DATA_BLOCK "DB_M256M_Scada"   // DB2011
{ S7_Optimized_Access := 'FALSE' }
VERSION : 0.1
   VAR
      tAlm : Struct   // HMI Alarms
         tE : Struct
            x0 : Bool;   // KE.Main emergency on
            x1 : Bool;   // KE1.Local emergency on
            x2 : Bool;   // Cabinet.Emergency localization
            x3 : Bool;   // SB1.Emergency localization
            x4 : Bool;   // SB2.Emergency localization
            x5 : Bool;
            x6 : Bool;
            x7 : Bool;
            x8 : Bool;
            x9 : Bool;
            x10 : Bool;
            x11 : Bool;
            x12 : Bool;
            x13 : Bool;
            x14 : Bool;
            x15 : Bool;
            x16 : Bool;
            x17 : Bool;
            x18 : Bool;
            x19 : Bool;
            x20 : Bool;
            x21 : Bool;
            x22 : Bool;
            x23 : Bool;
            x24 : Bool;
            x25 : Bool;
            x26 : Bool;
            x27 : Bool;
            x28 : Bool;
            x29 : Bool;
            x30 : Bool;
            x31 : Bool;
         END_STRUCT;
         tS : Struct
            tS0 : Struct
               x0 : Bool;   // xB18-3L+.PowerSupplyInputControlCabinetON / Head#1.Initialization timeout
               x1 : Bool;   // xB140QF2.ProtectionPowerSupplyMotorsYcut" / Head#1.homing timeout
               x2 : Bool;   // PLCA.Timeout receiving consumed message / Head#1.positioning timeout
               x3 : Bool;   // Syncro.Timeout receiving meter signal from main line / Head#1.carriage overload
               x4 : Bool;   // Head#1.drive error
               x5 : Bool;   // Head#1.missing ethernet IP connection
               x6 : Bool;   // Head#1.op.side overstroke
               x7 : Bool;   // Head#1.oppo.op.side overstroke
               x8 : Bool;   // Head#1.overstroke
               x9 : Bool;   // xB18-7L+.InputInstallationPowerSupplyON" / Head#2.Initialization timeout
               x10 : Bool;   // xB41QF2.Protection power supply motors longitudinal cutting / Head#2.homing timeout
               x11 : Bool;   // PLCB.Timeout receiving consumed message / Head#2.positioning timeout
               x12 : Bool;   // Syncro.Timeout receiving syncro value from mainline / Head#2.carriage overload
               x13 : Bool;   // Head#2.drive error
               x14 : Bool;   // Head#2.missing ethernet IP connection
               x15 : Bool;   // Head#2.op.side overstroke
               x16 : Bool;   // Head#2.oppo.op.side overstroke
               x17 : Bool;   // Head#2.overstroke
               x18 : Bool;   // xB11QF1/1D/QF2.Anomaly power supplies 120V / Head#3.Initialization timeout
               x19 : Bool;   // PLCA.Mission packet lost / Head#3.homing timeout
               x20 : Bool;   // Syncro.Unexpected syncro pulse / Head#3.positioning timeout
               x21 : Bool;   // Head#3.carriage overload
               x22 : Bool;   // Head#3.drive error
               x23 : Bool;   // Head#3.missing ethernet IP connection
               x24 : Bool;   // Head#3.op.side overstroke
               x25 : Bool;   // Head#3.oppo.op.side overstroke
               x26 : Bool;   // xB115KM1/2.AuxiliaryPowerSupplySetIn / Head#3.overstroke
               x27 : Bool;
               x28 : Bool;
               x29 : Bool;
               x30 : Bool;
               x31 : Bool;
            END_STRUCT;
            tS1 : Struct
               x0 : Bool;   // xB42QF2.Protection power supply motors longitudinal cutting / Head#4.Initialization timeout
               x1 : Bool;   // PLCB.Mission packet lost / Head#4.homing timeout
               x2 : Bool;   // Syncro.Unexpected syncro message / Head#4.positioning timeout
               x3 : Bool;   // Head#4.carriage overload
               x4 : Bool;   // Head#4.drive error
               x5 : Bool;   // Head#4.missing ethernet IP connection
               x6 : Bool;   // Head#4.op.side overstroke
               x7 : Bool;   // Head#4.oppo.op.side overstroke
               x8 : Bool;   // xB410AP1.SafetyOnPanel1" / Head#4.overstroke
               x9 : Bool;   // Head#5.Initialization timeout
               x10 : Bool;   // PLCA.Syncro packet lost / Head#5.homing timeout
               x11 : Bool;   // Syncro.Machine not syncronized / Head#5.positioning timeout
               x12 : Bool;   // Head#5.carriage overload
               x13 : Bool;   // Head#5.drive error
               x14 : Bool;   // Head#5.missing ethernet IP connection
               x15 : Bool;   // Head#5.op.side overstroke
               x16 : Bool;   // Head#5.oppo.op.side overstroke
               x17 : Bool;   // xB410AP1.SafetyOnPanel2" / Head#5.overstroke
               x18 : Bool;   // Head#6.Initialization timeout
               x19 : Bool;   // PLCB.Syncro packet lost / Head#6.homing timeout
               x20 : Bool;   // Head#6.positioning timeout
               x21 : Bool;   // Head#6.carriage overload
               x22 : Bool;   // Head#6.drive error
               x23 : Bool;   // Head#6.missing ethernet IP connection
               x24 : Bool;   // Head#6.op.side overstroke
               x25 : Bool;   // Head#6.oppo.op.side overstroke
               x26 : Bool;   // xB20QF3.Power supply 24V logic / Head#6.overstroke
               x27 : Bool;
               x28 : Bool;
               x29 : Bool;
               x30 : Bool;
               x31 : Bool;
            END_STRUCT;
            tS2 : Struct
               x0 : Bool;   // Head#7.Initialization timeout
               x1 : Bool;   // Syncro.YCut meter gap outside the limits / Head#7.homing timeout
               x2 : Bool;   // Head#7.positioning timeout
               x3 : Bool;   // Head#7.carriage overload
               x4 : Bool;   // Head#7.drive error
               x5 : Bool;   // Head#7.missing ethernet IP connection
               x6 : Bool;   // Head#7.op.side overstroke
               x7 : Bool;   // Head#7.oppo.op.side overstroke
               x8 : Bool;   // xB21QF1.Power supply 24V logic / Head#7.overstroke
               x9 : Bool;   // Head#8.Initialization timeout
               x10 : Bool;   // Syncro.Main line meter gap outside the limits / Head#8.homing timeout
               x11 : Bool;   // Head#8.positioning timeout
               x12 : Bool;   // Head#8.carriage overload
               x13 : Bool;   // Head#8.drive error
               x14 : Bool;   // Head#8.missing ethernet IP connection
               x15 : Bool;   // Head#8.op.side overstroke
               x16 : Bool;   // Head#8.oppo.op.side overstroke
               x17 : Bool;   // Head#8.overstroke
               x18 : Bool;
               x19 : Bool;
               x20 : Bool;
               x21 : Bool;
               x22 : Bool;
               x23 : Bool;
               x24 : Bool;
               x25 : Bool;
               x26 : Bool;
               x27 : Bool;
               x28 : Bool;
               x29 : Bool;
               x30 : Bool;
               x31 : Bool;
            END_STRUCT;
            tS3 : Struct
               x0 : Bool;
               x1 : Bool;   // Syncro.YCut meter gap outside the limits
               x2 : Bool;
               x3 : Bool;
               x4 : Bool;
               x5 : Bool;
               x6 : Bool;
               x7 : Bool;
               x8 : Bool;   // xB21QF1.Power supply 24V logic
               x9 : Bool;
               x10 : Bool;   // Syncro.Main line meter gap outside the limits
               x11 : Bool;
               x12 : Bool;
               x13 : Bool;
               x14 : Bool;
               x15 : Bool;
               x16 : Bool;
               x17 : Bool;
               x18 : Bool;
               x19 : Bool;
               x20 : Bool;
               x21 : Bool;
               x22 : Bool;
               x23 : Bool;
               x24 : Bool;
               x25 : Bool;
               x26 : Bool;
               x27 : Bool;
               x28 : Bool;
               x29 : Bool;
               x30 : Bool;
               x31 : Bool;
            END_STRUCT;
         END_STRUCT;
         tF : Struct
            x0 : Bool;
            x1 : Bool;
            x2 : Bool;
            x3 : Bool;
            x4 : Bool;
            x5 : Bool;
            x6 : Bool;
            x7 : Bool;
            x8 : Bool;
            x9 : Bool;
            x10 : Bool;
            x11 : Bool;
            x12 : Bool;
            x13 : Bool;
            x14 : Bool;
            x15 : Bool;
            x16 : Bool;
            x17 : Bool;
            x18 : Bool;
            x19 : Bool;
            x20 : Bool;
            x21 : Bool;
            x22 : Bool;
            x23 : Bool;
            x24 : Bool;
            x25 : Bool;
            x26 : Bool;
            x27 : Bool;
            x28 : Bool;
            x29 : Bool;
            x30 : Bool;
            x31 : Bool;
         END_STRUCT;
         tW : Struct
            x0 : Bool;   // PLCA.Timeout receiving consumed message
            x1 : Bool;   // PLCB.Timeout receiving consumed message
            x2 : Bool;   // PLCA.Mission packet lost
            x3 : Bool;   // PLCB.Mission packet lost
            x4 : Bool;   // PLCA.Syncro packet lost
            x5 : Bool;   // PLCB.Syncro packet lost
            x6 : Bool;   // QF.Protection air conditioners
            x7 : Bool;
            x8 : Bool;
            x9 : Bool;
            x10 : Bool;
            x11 : Bool;
            x12 : Bool;
            x13 : Bool;
            x14 : Bool;
            x15 : Bool;
            x16 : Bool;
            x17 : Bool;
            x18 : Bool;
            x19 : Bool;
            x20 : Bool;
            x21 : Bool;
            x22 : Bool;
            x23 : Bool;
            x24 : Bool;
            x25 : Bool;
            x26 : Bool;
            x27 : Bool;
            x28 : Bool;
            x29 : Bool;
            x30 : Bool;
            x31 : Bool;
         END_STRUCT;
      END_STRUCT;
      tHMR : Struct   // HMI Read
         xSpare0 : Bool := FALSE;   // Calibration function allowed {x|x|x|x|O}
         xSpare1 : Bool;
         xSpare2 : Bool;
         xSpare3 : Bool;
         xSpare4 : Bool;
         xSpare5 : Bool;
         xSpare6 : Bool;
         xSpare7 : Bool;
         xSpare8 : Bool;
         xSpare9 : Bool;
         xSpare10 : Bool;
         xSpare11 : Bool;
         xSpare12 : Bool;
         xSpare13 : Bool;
         xSpare14 : Bool;
         xSpare15 : Bool := FALSE;
         xSpare16 : Bool;
         xSpare17 : Bool;
         xSpare18 : Bool;
         xSpare19 : Bool;
         xSpare20 : Bool;
         xSpare21 : Bool;
         xSpare22 : Bool;
         xSpare23 : Bool;
         xSpare24 : Bool;
         xSpare25 : Bool;
         xSpare26 : Bool;
         xSpare27 : Bool;
         xSpare28 : Bool;
         xSpare29 : Bool;
         xSpare30 : Bool;
         xSpare31 : Bool;
         xSpare : Array[0..15] of Bool;
         iCodeAlarm_H1 : Int;   // Motor error code H1
         iCodeAlarm_H2 : Int;   // Motor error code H2
         iCodeAlarm_H3 : Int;   // Motor error code H3
         iCodeAlarm_H4 : Int;   // Motor error code H4
         iCodeAlarm_H5 : Int;   // Motor error code H5
         iCodeAlarm_H6 : Int;   // Motor error code H6
         iCodeAlarm_H7 : Int;   // Motor error code H7
         iCodeAlarm_H8 : Int;   // Motor error code H8
         iSpare8 : Int;
         iSpare9 : Int;
         iSpare10 : Int;
         iSpare11 : Int;
         iSpare12 : Int;
         iSpare13 : Int;
         iSpare14 : Int;
         iSpare15 : Int;
         iSpare16 : Int;
         dHeadActualPositions_cmm_H1 : DInt;   // Head#x head actual position [mm/100] {mm/100|mm|x|x|O} / Head#1 head actual position [mm/100] {mm/100|mm|x|x|O}
         dHeadActualPositions_cmm_H2 : DInt;   // Head#x head actual position [mm/100] {mm/100|mm|x|x|O} / Head#2 head actual position [mm/100] {mm/100|mm|x|x|O}
         dHeadActualPositions_cmm_H3 : DInt;   // Head#x head actual position [mm/100] {mm/100|mm|x|x|O} / Head#3 head actual position [mm/100] {mm/100|mm|x|x|O}
         dHeadActualPositions_cmm_H4 : DInt;   // Head#x head actual position [mm/100] {mm/100|mm|x|x|O} / Head#4 head actual position [mm/100] {mm/100|mm|x|x|O}
         dHeadActualPositions_cmm_H5 : DInt;   // Head#x head actual position [mm/100] {mm/100|mm|x|x|O} / Head#5 head actual position [mm/100] {mm/100|mm|x|x|O}
         dHeadActualPositions_cmm_H6 : DInt;   // Head#x head actual position [mm/100] {mm/100|mm|x|x|O} / Head#6 head actual position [mm/100] {mm/100|mm|x|x|O}
         dHeadActualPositions_cmm_H7 : DInt;   // Head#x head actual position [mm/100] {mm/100|mm|x|x|O} / Head#7 head actual position [mm/100] {mm/100|mm|x|x|O}
         dHeadActualPositions_cmm_H8 : DInt;   // Head#x head actual position [mm/100] {mm/100|mm|x|x|O} / Head#8 head actual position [mm/100] {mm/100|mm|x|x|O}
         dHeadHomePositions_cmm_H1 : DInt;   // Head#x home position [mm/100] {mm/100|mm|x|x|O} / Head#1 home position [mm/100] {mm/100|mm|x|x|O}
         dHeadHomePositions_cmm_H2 : DInt;   // Head#x home position [mm/100] {mm/100|mm|x|x|O} / Head#2 home position [mm/100] {mm/100|mm|x|x|O}
         dHeadHomePositions_cmm_H3 : DInt;   // Head#x home position [mm/100] {mm/100|mm|x|x|O} / Head#3 home position [mm/100] {mm/100|mm|x|x|O}
         dHeadHomePositions_cmm_H4 : DInt;   // Head#x home position [mm/100] {mm/100|mm|x|x|O} / Head#4 home position [mm/100] {mm/100|mm|x|x|O}
         dHeadHomePositions_cmm_H5 : DInt;   // Head#x home position [mm/100] {mm/100|mm|x|x|O} / Head#5 home position [mm/100] {mm/100|mm|x|x|O}
         dHeadHomePositions_cmm_H6 : DInt;   // Head#x home position [mm/100] {mm/100|mm|x|x|O} / Head#6 home position [mm/100] {mm/100|mm|x|x|O}
         dHeadHomePositions_cmm_H7 : DInt;   // Head#x home position [mm/100] {mm/100|mm|x|x|O} / Head#7 home position [mm/100] {mm/100|mm|x|x|O}
         dHeadHomePositions_cmm_H8 : DInt;   // Head#x home position [mm/100] {mm/100|mm|x|x|O} / Head#8 home position [mm/100] {mm/100|mm|x|x|O}
         dHeadMoveStatus_H1 : DInt;   // Head#x move status (1=Not Initialized 2=Not referred 3=Not positioned 4=Positioned 5=Positioning 6=Virtual collision 7=Anomaly) {x|x|x|x|O} / Head#1 move status (1=Not Initialized 2=Not referred 3=Not positioned 4=Positioned 5=Positioning 6=Virtual collision 7=Anomaly) {x|x|x|x|O}
         dHeadMoveStatus_H2 : DInt;   // Head#x move status (1=Not Initialized 2=Not referred 3=Not positioned 4=Positioned 5=Positioning 6=Virtual collision 7=Anomaly) {x|x|x|x|O} / Head#2 move status (1=Not Initialized 2=Not referred 3=Not positioned 4=Positioned 5=Positioning 6=Virtual collision 7=Anomaly) {x|x|x|x|O}
         dHeadMoveStatus_H3 : DInt;   // Head#x move status (1=Not Initialized 2=Not referred 3=Not positioned 4=Positioned 5=Positioning 6=Virtual collision 7=Anomaly) {x|x|x|x|O} / Head#3 move status (1=Not Initialized 2=Not referred 3=Not positioned 4=Positioned 5=Positioning 6=Virtual collision 7=Anomaly) {x|x|x|x|O}
         dHeadMoveStatus_H4 : DInt;   // Head#x move status (1=Not Initialized 2=Not referred 3=Not positioned 4=Positioned 5=Positioning 6=Virtual collision 7=Anomaly) {x|x|x|x|O} / Head#4 move status (1=Not Initialized 2=Not referred 3=Not positioned 4=Positioned 5=Positioning 6=Virtual collision 7=Anomaly) {x|x|x|x|O}
         dHeadMoveStatus_H5 : DInt;   // Head#x move status (1=Not Initialized 2=Not referred 3=Not positioned 4=Positioned 5=Positioning 6=Virtual collision 7=Anomaly) {x|x|x|x|O} / Head#5 move status (1=Not Initialized 2=Not referred 3=Not positioned 4=Positioned 5=Positioning 6=Virtual collision 7=Anomaly) {x|x|x|x|O}
         dHeadMoveStatus_H6 : DInt;   // Head#x move status (1=Not Initialized 2=Not referred 3=Not positioned 4=Positioned 5=Positioning 6=Virtual collision 7=Anomaly) {x|x|x|x|O} / Head#6 move status (1=Not Initialized 2=Not referred 3=Not positioned 4=Positioned 5=Positioning 6=Virtual collision 7=Anomaly) {x|x|x|x|O}
         dHeadMoveStatus_H7 : DInt;   // Head#x move status (1=Not Initialized 2=Not referred 3=Not positioned 4=Positioned 5=Positioning 6=Virtual collision 7=Anomaly) {x|x|x|x|O} / Head#7 move status (1=Not Initialized 2=Not referred 3=Not positioned 4=Positioned 5=Positioning 6=Virtual collision 7=Anomaly) {x|x|x|x|O}
         dHeadMoveStatus_H8 : DInt;   // Head#x move status (1=Not Initialized 2=Not referred 3=Not positioned 4=Positioned 5=Positioning 6=Virtual collision 7=Anomaly) {x|x|x|x|O} / Head#8 move status (1=Not Initialized 2=Not referred 3=Not positioned 4=Positioned 5=Positioning 6=Virtual collision 7=Anomaly) {x|x|x|x|O}
         dSpare : Array[0..7] of DInt;
         rSpare0 : Real;
         rSpare1 : Real;
         rSpare2 : Real;
         rSpare3 : Real;
         rSpare4 : Real;
         rSpare5 : Real;
         rSpare6 : Real;
         rSpare7 : Real;
         rSpare8 : Real;
         tManCmd : Struct
            xManJogForwardFdbk_H1 : Bool;   // Head#x manual jog forward fdbk {x|x|x|x|O} / Head#1 manual jog forward fdbk {x|x|x|x|O}
            xManJogBackwardFdbk_H1 : Bool;   // Head#x manual jog backward fdbk {x|x|x|x|O} / Head#1 manual jog backward fdbk {x|x|x|x|O}
            xManJogForwardFdbk_H2 : Bool;   // Head#x manual jog forward fdbk {x|x|x|x|O} / Head#2 manual jog forward fdbk {x|x|x|x|O}
            xManJogBackwardFdbk_H2 : Bool;   // Head#x manual jog backward fdbk {x|x|x|x|O} / Head#2 manual jog backward fdbk {x|x|x|x|O}
            xManJogForwardFdbk_H3 : Bool;   // Head#x manual jog forward fdbk {x|x|x|x|O} / Head#3 manual jog forward fdbk {x|x|x|x|O}
            xManJogBackwardFdbk_H3 : Bool;   // Head#x manual jog backward fdbk {x|x|x|x|O} / Head#3 manual jog backward fdbk {x|x|x|x|O}
            xManJogForwardFdbk_H4 : Bool;   // Head#x manual jog forward fdbk {x|x|x|x|O} / Head#4 manual jog forward fdbk {x|x|x|x|O}
            xManJogBackwardFdbk_H4 : Bool;   // Head#x manual jog backward fdbk {x|x|x|x|O} / Head#4 manual jog backward fdbk {x|x|x|x|O}
            xManJogForwardFdbk_H5 : Bool;   // Head#x manual jog forward fdbk {x|x|x|x|O} / Head#5 manual jog forward fdbk {x|x|x|x|O}
            xManJogBackwardFdbk_H5 : Bool;   // Head#x manual jog backward fdbk {x|x|x|x|O} / Head#5 manual jog backward fdbk {x|x|x|x|O}
            xManJogForwardFdbk_H6 : Bool;   // Head#x manual jog forward fdbk {x|x|x|x|O} / Head#6 manual jog forward fdbk {x|x|x|x|O}
            xManJogBackwardFdbk_H6 : Bool;   // Head#x manual jog backward fdbk {x|x|x|x|O} / Head#6 manual jog backward fdbk {x|x|x|x|O}
            xManJogForwardFdbk_H7 : Bool;   // Head#x manual jog forward fdbk {x|x|x|x|O} / Head#7 manual jog forward fdbk {x|x|x|x|O}
            xManJogBackwardFdbk_H7 : Bool;   // Head#x manual jog backward fdbk {x|x|x|x|O} / Head#7 manual jog backward fdbk {x|x|x|x|O}
            xManJogForwardFdbk_H8 : Bool;   // Head#x manual jog forward fdbk {x|x|x|x|O} / Head#8 manual jog forward fdbk {x|x|x|x|O}
            xManJogBackwardFdbk_H8 : Bool;   // Head#x manual jog backward fdbk {x|x|x|x|O} / Head#8 manual jog backward fdbk {x|x|x|x|O}
            xSpare : Array[0..15] of Bool;
         END_STRUCT;
      END_STRUCT;
      tHMW : Struct   // HMI Write
         xBrakeRealeaseHead_H1 : Bool := FALSE;   // Force the brake release of the head {x|x|x|x|M} / Force the brake release of the Head #1 {x|x|x|x|M}
         xBrakeEngageHeads_H1 : Bool := FALSE;   // Force the brake engaged of the head {x|x|x|x|M} / Force the brake engaged of the Head #1 {x|x|x|x|M}
         xUpdateHomeHead_H1 : Bool;   // Update home position head#x {x|x|x|x|M} / Update home position Head #1 {x|x|x|x|M}
         xBrakeRealeaseHead_H2 : Bool := FALSE;   // Force the brake release of the head {x|x|x|x|M} / Force the brake release of the Head #2 {x|x|x|x|M}
         xBrakeEngageHeads_H2 : Bool := FALSE;   // Force the brake engaged of the head {x|x|x|x|M} / Force the brake engaged of the Head #2 {x|x|x|x|M}
         xUpdateHomeHead_H2 : Bool;   // Update home position head#x {x|x|x|x|M} / Update home position Head #2 {x|x|x|x|M}
         xBrakeRealeaseHead_H3 : Bool := FALSE;   // Force the brake release of the head {x|x|x|x|M} / Force the brake release of the Head #3 {x|x|x|x|M}
         xBrakeEngageHeads_H3 : Bool := FALSE;   // Force the brake engaged of the head {x|x|x|x|M} / Force the brake engaged of the Head #3 {x|x|x|x|M}
         xUpdateHomeHead_H3 : Bool;   // Update home position head#x {x|x|x|x|M} / Update home position Head #3 {x|x|x|x|M}
         xBrakeRealeaseHead_H4 : Bool := FALSE;   // Force the brake release of the head {x|x|x|x|M} / Force the brake release of the Head #4{x|x|x|x|M}
         xBrakeEngageHeads_H4 : Bool := FALSE;   // Force the brake engaged of the head {x|x|x|x|M} / Force the brake engaged of the Head #4{x|x|x|x|M}
         xUpdateHomeHead_H4 : Bool;   // Update home position head#x {x|x|x|x|M} / Update home position Head #4 {x|x|x|x|M}
         xBrakeRealeaseHead_H5 : Bool := FALSE;   // Force the brake release of the head {x|x|x|x|M} / Force the brake release of the Head #5{x|x|x|x|M}
         xBrakeEngageHeads_H5 : Bool := FALSE;   // Force the brake engaged of the head {x|x|x|x|M} / Force the brake engaged of the Head #5{x|x|x|x|M}
         xUpdateHomeHead_H5 : Bool;   // Update home position head#x {x|x|x|x|M} / Update home position Head #5 {x|x|x|x|M}
         xBrakeRealeaseHead_H6 : Bool := FALSE;   // Force the brake release of the head {x|x|x|x|M} / Force the brake release of the Head #6{x|x|x|x|M}
         xBrakeEngageHeads_H6 : Bool := FALSE;   // Force the brake engaged of the head {x|x|x|x|M} / Force the brake engaged of the Head #6 {x|x|x|x|M}
         xUpdateHomeHead_H6 : Bool;   // Update home position head#x {x|x|x|x|M} / Update home position Head #6 {x|x|x|x|M}
         xBrakeRealeaseHead_H7 : Bool := FALSE;   // Force the brake release of the head {x|x|x|x|M} / Force the brake release of the Head #7{x|x|x|x|M}
         xBrakeEngageHeads_H7 : Bool := FALSE;   // Force the brake engaged of the head {x|x|x|x|M} / Force the brake engaged of the Head #7{x|x|x|x|M}
         xUpdateHomeHead_H7 : Bool;   // Update home position head#x {x|x|x|x|M} / Update home position Head #7{x|x|x|x|M}
         xBrakeRealeaseHead_H8 : Bool := FALSE;   // Force the brake release of the head {x|x|x|x|M} / Force the brake release of the Head #8{x|x|x|x|M}
         xBrakeEngageHeads_H8 : Bool := FALSE;   // Force the brake engaged of the head {x|x|x|x|M} / Force the brake engaged of the Head #8{x|x|x|x|M}
         xUpdateHomeHead_H8 : Bool;   // Update home position head#x {x|x|x|x|M} / Update home position Head #8 {x|x|x|x|M}
         xSpare24 : Bool;
         xSpare25 : Bool;
         xSpare26 : Bool;
         xSpare27 : Bool;
         xSpare28 : Bool;
         xSpare29 : Bool;
         xSpare30 : Bool;
         xSpare31 : Bool;
         xSpare : Array[0..15] of Bool;
         iSpare0 : Int;
         iSpare1 : Int;
         iSpare2 : Int;
         iSpare3 : Int;
         iSpare4 : Int;
         iSpare5 : Int;
         iSpare6 : Int;
         iSpare7 : Int;
         iSpare8 : Int;
         iSpare9 : Int;
         iSpare10 : Int;
         iSpare11 : Int;
         iSpare12 : Int;
         iSpare13 : Int;
         iSpare14 : Int;
         iSpare15 : Int;
         iSpare16 : Int;
         dHeadHomePositions_cmm_H1 : DInt;   // Head#x home position [mm/100] {mm/100|mm|-2500|2500|M} / Head#1 home position [mm/100] {mm/100|mm|-2500|2500|M}
         dHeadHomePositions_cmm_H2 : DInt;   // Head#x home position [mm/100] {mm/100|mm|-2500|2500|M} / Head#2 home position [mm/100] {mm/100|mm|-2500|2500|M}
         dHeadHomePositions_cmm_H3 : DInt;   // Head#x home position [mm/100] {mm/100|mm|-2500|2500|M} / Head#3 home position [mm/100] {mm/100|mm|-2500|2500|M}
         dHeadHomePositions_cmm_H4 : DInt;   // Head#x home position [mm/100] {mm/100|mm|-2500|2500|M} / Head#4 home position [mm/100] {mm/100|mm|-2500|2500|M}
         dHeadHomePositions_cmm_H5 : DInt;   // Head#x home position [mm/100] {mm/100|mm|-2500|2500|M} / Head#5 home position [mm/100] {mm/100|mm|-2500|2500|M}
         dHeadHomePositions_cmm_H6 : DInt;   // Head#x home position [mm/100] {mm/100|mm|-2500|2500|M} / Head#6 home position [mm/100] {mm/100|mm|-2500|2500|M}
         dHeadHomePositions_cmm_H7 : DInt;   // Head#x home position [mm/100] {mm/100|mm|-2500|2500|M} / Head#7 home position [mm/100] {mm/100|mm|-2500|2500|M}
         dHeadHomePositions_cmm_H8 : DInt;   // Head#x home position [mm/100] {mm/100|mm|-2500|2500|M} / Head#8 home position [mm/100] {mm/100|mm|-2500|2500|M}
         dSpare8 : DInt;
         dSpare9 : DInt;
         dSpare10 : DInt;
         dSpare11 : DInt;
         dSpare12 : DInt;
         dSpare13 : DInt;
         dSpare14 : DInt;
         dSpare15 : DInt;
         dSpare : Array[0..43] of DInt;
         rSpare0 : Real;
         rSpare1 : Real;
         rSpare2 : Real;
         rSpare3 : Real;
         rSpare4 : Real;
         rSpare5 : Real;
         rSpare6 : Real;
         rSpare7 : Real;
         rSpare8 : Real;
         tManCmd : Struct
            xMan_JogForward_H1 : Bool;   // Head #x manual jog forward {x|x|x|x|O} / Head #1 manual jog forward {x|x|x|x|O}
            xMan_JogBackward_H1 : Bool;   // Head #x manual jog backward {x|x|x|x|O} / Head #1 manual jog backward {x|x|x|x|O}
            xMan_JogForward_H2 : Bool;   // Head #x manual jog forward {x|x|x|x|O} / Head #2 manual jog forward {x|x|x|x|O}
            xMan_JogBackward_H2 : Bool;   // Head #x manual jog backward {x|x|x|x|O} / Head #2 manual jog backward {x|x|x|x|O}
            xMan_JogForward_H3 : Bool;   // Head #x manual jog forward {x|x|x|x|O} / Head #3 manual jog forward {x|x|x|x|O}
            xMan_JogBackward_H3 : Bool;   // Head #x manual jog backward {x|x|x|x|O} / Head #3 manual jog backward {x|x|x|x|O}
            xMan_JogForward_H4 : Bool;   // Head #x manual jog forward {x|x|x|x|O} / Head #4 manual jog forward {x|x|x|x|O}
            xMan_JogBackward_H4 : Bool;   // Head #x manual jog backward {x|x|x|x|O} / Head #4 manual jog backward {x|x|x|x|O}
            xMan_JogForward_H5 : Bool;   // Head #x manual jog forward {x|x|x|x|O} / Head #5 manual jog forward {x|x|x|x|O}
            xMan_JogBackward_H5 : Bool;   // Head #x manual jog backward {x|x|x|x|O} / Head #5 manual jog backward {x|x|x|x|O}
            xMan_JogForward_H6 : Bool;   // Head #x manual jog forward {x|x|x|x|O} / Head #6 manual jog forward {x|x|x|x|O}
            xMan_JogBackward_H6 : Bool;   // Head #x manual jog backward {x|x|x|x|O} / Head #6 manual jog backward {x|x|x|x|O}
            xMan_JogForward_H7 : Bool;   // Head #x manual jog forward {x|x|x|x|O} / Head #7 manual jog forward {x|x|x|x|O}
            xMan_JogBackward_H7 : Bool;   // Head #x manual jog backward {x|x|x|x|O} / Head #7 manual jog backward {x|x|x|x|O}
            xMan_JogForward_H8 : Bool;   // Head #x manual jog forward {x|x|x|x|O} / Head #8 manual jog forward {x|x|x|x|O}
            xMan_JogBackward_H8 : Bool;   // Head #x manual jog backward {x|x|x|x|O} / Head #8 manual jog backward {x|x|x|x|O}
            xSpare16 : Bool;
            xSpare17 : Bool;
            xSpare18 : Bool;
            xSpare19 : Bool;
            xSpare20 : Bool;
            xSpare21 : Bool;
            xSpare22 : Bool;
            xSpare23 : Bool;
            xSpare24 : Bool;
            xSpare25 : Bool;
            xSpare26 : Bool;
            xSpare27 : Bool;
            xSpare28 : Bool;
            xSpare29 : Bool;
            xSpare30 : Bool;
            xSpare31 : Bool;
         END_STRUCT;
      END_STRUCT;
   END_VAR
BEGIN
END_DATA_BLOCK

DATA_BLOCK "DB_M256F_Scada"   // DB2012
{ S7_Optimized_Access := 'FALSE' }
VERSION : 0.1
   VAR
      tAlm : Struct   // HMI Alarms
         tE : Struct
            x0 : Bool;   // KE.Main emergency on
            x1 : Bool;   // KE1.Local emergency on
            x2 : Bool;   // Cabinet.Emergency localization
            x3 : Bool;   // SB1.Emergency localization
            x4 : Bool;   // SB2.Emergency localization
            x5 : Bool;
            x6 : Bool;
            x7 : Bool;
            x8 : Bool;
            x9 : Bool;
            x10 : Bool;
            x11 : Bool;
            x12 : Bool;
            x13 : Bool;
            x14 : Bool;
            x15 : Bool;
            x16 : Bool;
            x17 : Bool;
            x18 : Bool;
            x19 : Bool;
            x20 : Bool;
            x21 : Bool;
            x22 : Bool;
            x23 : Bool;
            x24 : Bool;
            x25 : Bool;
            x26 : Bool;
            x27 : Bool;
            x28 : Bool;
            x29 : Bool;
            x30 : Bool;
            x31 : Bool;
         END_STRUCT;
         tS : Struct
            tS0 : Struct
               x0 : Bool;
               x1 : Bool;   // Syncro.YCut meter gap outside the limits
               x2 : Bool;
               x3 : Bool;
               x4 : Bool;
               x5 : Bool;
               x6 : Bool;
               x7 : Bool;
               x8 : Bool;   // xB21QF1.Power supply 24V logic
               x9 : Bool;
               x10 : Bool;   // Syncro.Main line meter gap outside the limits
               x11 : Bool;
               x12 : Bool;
               x13 : Bool;
               x14 : Bool;
               x15 : Bool;
               x16 : Bool;
               x17 : Bool;
               x18 : Bool;
               x19 : Bool;
               x20 : Bool;
               x21 : Bool;
               x22 : Bool;
               x23 : Bool;
               x24 : Bool;
               x25 : Bool;
               x26 : Bool;
               x27 : Bool;
               x28 : Bool;
               x29 : Bool;
               x30 : Bool;
               x31 : Bool;
            END_STRUCT;
            tS1 : Struct
               x0 : Bool;
               x1 : Bool;   // Syncro.YCut meter gap outside the limits
               x2 : Bool;
               x3 : Bool;
               x4 : Bool;
               x5 : Bool;
               x6 : Bool;
               x7 : Bool;
               x8 : Bool;   // xB21QF1.Power supply 24V logic
               x9 : Bool;
               x10 : Bool;   // Syncro.Main line meter gap outside the limits
               x11 : Bool;
               x12 : Bool;
               x13 : Bool;
               x14 : Bool;
               x15 : Bool;
               x16 : Bool;
               x17 : Bool;
               x18 : Bool;
               x19 : Bool;
               x20 : Bool;
               x21 : Bool;
               x22 : Bool;
               x23 : Bool;
               x24 : Bool;
               x25 : Bool;
               x26 : Bool;
               x27 : Bool;
               x28 : Bool;
               x29 : Bool;
               x30 : Bool;
               x31 : Bool;
            END_STRUCT;
            tS2 : Struct
               x0 : Bool;
               x1 : Bool;   // Syncro.YCut meter gap outside the limits
               x2 : Bool;
               x3 : Bool;
               x4 : Bool;
               x5 : Bool;
               x6 : Bool;
               x7 : Bool;
               x8 : Bool;   // xB21QF1.Power supply 24V logic
               x9 : Bool;
               x10 : Bool;   // Syncro.Main line meter gap outside the limits
               x11 : Bool;
               x12 : Bool;
               x13 : Bool;
               x14 : Bool;
               x15 : Bool;
               x16 : Bool;
               x17 : Bool;
               x18 : Bool;
               x19 : Bool;
               x20 : Bool;
               x21 : Bool;
               x22 : Bool;
               x23 : Bool;
               x24 : Bool;
               x25 : Bool;
               x26 : Bool;
               x27 : Bool;
               x28 : Bool;
               x29 : Bool;
               x30 : Bool;
               x31 : Bool;
            END_STRUCT;
            tS3 : Struct
               x0 : Bool;
               x1 : Bool;   // Syncro.YCut meter gap outside the limits
               x2 : Bool;
               x3 : Bool;
               x4 : Bool;
               x5 : Bool;
               x6 : Bool;
               x7 : Bool;
               x8 : Bool;   // xB21QF1.Power supply 24V logic
               x9 : Bool;
               x10 : Bool;   // Syncro.Main line meter gap outside the limits
               x11 : Bool;
               x12 : Bool;
               x13 : Bool;
               x14 : Bool;
               x15 : Bool;
               x16 : Bool;
               x17 : Bool;
               x18 : Bool;
               x19 : Bool;
               x20 : Bool;
               x21 : Bool;
               x22 : Bool;
               x23 : Bool;
               x24 : Bool;
               x25 : Bool;
               x26 : Bool;
               x27 : Bool;
               x28 : Bool;
               x29 : Bool;
               x30 : Bool;
               x31 : Bool;
            END_STRUCT;
         END_STRUCT;
         tF : Struct
            x0 : Bool;
            x1 : Bool;
            x2 : Bool;
            x3 : Bool;
            x4 : Bool;
            x5 : Bool;
            x6 : Bool;
            x7 : Bool;
            x8 : Bool;
            x9 : Bool;
            x10 : Bool;
            x11 : Bool;
            x12 : Bool;
            x13 : Bool;
            x14 : Bool;
            x15 : Bool;
            x16 : Bool;
            x17 : Bool;
            x18 : Bool;
            x19 : Bool;
            x20 : Bool;
            x21 : Bool;
            x22 : Bool;
            x23 : Bool;
            x24 : Bool;
            x25 : Bool;
            x26 : Bool;
            x27 : Bool;
            x28 : Bool;
            x29 : Bool;
            x30 : Bool;
            x31 : Bool;
         END_STRUCT;
         tW : Struct
            x0 : Bool;   // PLCA.Timeout receiving consumed message
            x1 : Bool;   // PLCB.Timeout receiving consumed message
            x2 : Bool;   // PLCA.Mission packet lost
            x3 : Bool;   // PLCB.Mission packet lost
            x4 : Bool;   // PLCA.Syncro packet lost
            x5 : Bool;   // PLCB.Syncro packet lost
            x6 : Bool;   // QF.Protection air conditioners
            x7 : Bool;
            x8 : Bool;
            x9 : Bool;
            x10 : Bool;
            x11 : Bool;
            x12 : Bool;
            x13 : Bool;
            x14 : Bool;
            x15 : Bool;
            x16 : Bool;
            x17 : Bool;
            x18 : Bool;
            x19 : Bool;
            x20 : Bool;
            x21 : Bool;
            x22 : Bool;
            x23 : Bool;
            x24 : Bool;
            x25 : Bool;
            x26 : Bool;
            x27 : Bool;
            x28 : Bool;
            x29 : Bool;
            x30 : Bool;
            x31 : Bool;
         END_STRUCT;
      END_STRUCT;
      tHMR : Struct   // HMI Read
         xSpare0 : Bool;
         xSpare1 : Bool;
         xSpare2 : Bool;
         xSpare3 : Bool;
         xSpare4 : Bool;
         xSpare5 : Bool;
         xSpare6 : Bool;
         xSpare7 : Bool;
         xSpare8 : Bool;
         xSpare9 : Bool;
         xSpare10 : Bool;
         xSpare11 : Bool;
         xSpare12 : Bool;
         xSpare13 : Bool;
         xSpare14 : Bool;
         xSpare15 : Bool := FALSE;
         xSpare16 : Bool;
         xSpare17 : Bool;
         xSpare18 : Bool;
         xSpare19 : Bool;
         xSpare20 : Bool;
         xSpare21 : Bool;
         xSpare22 : Bool;
         xSpare23 : Bool;
         xSpare24 : Bool;
         xSpare25 : Bool;
         xSpare26 : Bool;
         xSpare27 : Bool;
         xSpare28 : Bool;
         xSpare29 : Bool;
         xSpare30 : Bool;
         xSpare31 : Bool;
         xSpare : Array[0..15] of Bool;
         iSpare0 : Int;
         iSpare1 : Int;
         iSpare2 : Int;
         iSpare3 : Int;
         iSpare4 : Int;
         iSpare5 : Int;
         iSpare6 : Int;
         iSpare7 : Int;
         iSpare8 : Int;
         iSpare9 : Int;
         iSpare10 : Int;
         iSpare11 : Int;
         iSpare12 : Int;
         iSpare13 : Int;
         iSpare14 : Int;
         iSpare15 : Int;
         iSpare16 : Int;
         dHeadStatus_H1 : DInt;   // Head#x firing status (1=OFF 3=ON) {x|x|x|x|O} / Head #1 firing status (1=OFF 3=ON) {x|x|x|x|O}
         dHeadStatus_H2 : DInt;   // Head#x firing status (1=OFF 3=ON) {x|x|x|x|O} / Head #2 firing status (1=OFF 3=ON) {x|x|x|x|O}
         dHeadStatus_H3 : DInt;   // Head#x firing status (1=OFF 3=ON) {x|x|x|x|O} / Head #3 firing status (1=OFF 3=ON) {x|x|x|x|O}
         dHeadStatus_H4 : DInt;   // Head#x firing status (1=OFF 3=ON) {x|x|x|x|O} / Head #4 firing status (1=OFF 3=ON) {x|x|x|x|O}
         dHeadStatus_H5 : DInt;   // Head#x firing status (1=OFF 3=ON) {x|x|x|x|O} / Head #5 firing status (1=OFF 3=ON) {x|x|x|x|O}
         dHeadStatus_H6 : DInt;   // Head#x firing status (1=OFF 3=ON) {x|x|x|x|O} / Head #6 firing status (1=OFF 3=ON) {x|x|x|x|O}
         dHeadStatus_H7 : DInt;   // Head#x firing status (1=OFF 3=ON) {x|x|x|x|O} / Head #7 firing status (1=OFF 3=ON) {x|x|x|x|O}
         dHeadStatus_H8 : DInt;   // Head#x firing status (1=OFF 3=ON) {x|x|x|x|O} / Head #8 firing status (1=OFF 3=ON) {x|x|x|x|O}
         dSpare8 : DInt := 0;
         dSpare9 : DInt := 0;
         dSpare10 : DInt := 0;
         dSpare11 : DInt := 0;
         dSpare12 : DInt;
         dSpare13 : DInt;
         dSpare14 : DInt;
         dSpare15 : DInt;
         dSpare : Array[0..15] of DInt;
         rHeadUsage_km_H1 : Real;   // Head#x head usage [km] {km|km|x|x|O} / Head #1 head usage [km] {km|km|x|x|O}
         rHeadUsage_km_H2 : Real;   // Head#x head usage [km] {km|km|x|x|O} / Head #2 head usage [km] {km|km|x|x|O}
         rHeadUsage_km_H3 : Real;   // Head#x head usage [km] {km|km|x|x|O} / Head #3 head usage [km] {km|km|x|x|O}
         rHeadUsage_km_H4 : Real;   // Head#x head usage [km] {km|km|x|x|O} / Head #4 head usage [km] {km|km|x|x|O}
         rHeadUsage_km_H5 : Real;   // Head#x head usage [km] {km|km|x|x|O} / Head #5 head usage [km] {km|km|x|x|O}
         rHeadUsage_km_H6 : Real;   // Head#x head usage [km] {km|km|x|x|O} / Head #6 head usage [km] {km|km|x|x|O}
         rHeadUsage_km_H7 : Real;   // Head#x head usage [km] {km|km|x|x|O} / Head #7 head usage [km] {km|km|x|x|O}
         rHeadUsage_km_H8 : Real;   // Head#x head usage [km] {km|km|x|x|O} / Head #8 head usage [km] {km|km|x|x|O}
         rSpare8 : Real;
         tManCmd : Struct
            xMan_FireON_Fdbk_H1 : Bool;   // Head#x manual fire ON Feeback {x|x|x|x|O} / Head #1 manual fire ON Feeback {x|x|x|x|O}
            xMan_FireOFF_Fdbk_H1 : Bool;   // Head#x manual fire OFF Feedback {x|x|x|x|O} / Head #1 manual fire OFF Feedback {x|x|x|x|O}
            xMan_OilON_Fdbk_H1 : Bool;   // Head#x manual oil feedback ON {x|x|x|x|O} / Head #1 manual oil feedback ON {x|x|x|x|O}
            xMan_FireON_Fdbk_H2 : Bool;   // Head#x manual fire ON Feeback {x|x|x|x|O} / Head #2 manual fire ON Feeback {x|x|x|x|O}
            xMan_FireOFF_Fdbk_H2 : Bool;   // Head#x manual fire OFF Feedback {x|x|x|x|O} / Head #2 manual fire OFF Feedback {x|x|x|x|O}
            xMan_OilON_Fdbk_H2 : Bool;   // Head#x manual oil feedback ON {x|x|x|x|O} / Head #2 manual oil feedback ON {x|x|x|x|O}
            xMan_FireON_Fdbk_H3 : Bool;   // Head#x manual fire ON Feeback {x|x|x|x|O} / Head #3 manual fire ON Feeback {x|x|x|x|O}
            xMan_FireOFF_Fdbk_H3 : Bool;   // Head#x manual fire OFF Feedback {x|x|x|x|O} / Head #3 manual fire OFF Feedback {x|x|x|x|O}
            xMan_OilON_Fdbk_H3 : Bool;   // Head#x manual oil feedback ON {x|x|x|x|O} / Head #3 manual oil feedback ON {x|x|x|x|O}
            xMan_FireON_Fdbk_H4 : Bool;   // Head#x manual fire ON Feeback {x|x|x|x|O} / Head #4 manual fire ON Feeback {x|x|x|x|O}
            xMan_FireOFF_Fdbk_H4 : Bool;   // Head#x manual fire OFF Feedback {x|x|x|x|O} / Head #4 manual fire OFF Feedback {x|x|x|x|O}
            xMan_OilON_Fdbk_H4 : Bool;   // Head#x manual oil feedback ON {x|x|x|x|O} / Head #4 manual oil feedback ON {x|x|x|x|O}
            xMan_FireON_Fdbk_H5 : Bool;   // Head#x manual fire ON Feeback {x|x|x|x|O} / Head #5 manual fire ON Feeback {x|x|x|x|O}
            xMan_FireOFF_Fdbk_H5 : Bool;   // Head#x manual fire OFF Feedback {x|x|x|x|O} / Head #5 manual fire OFF Feedback {x|x|x|x|O}
            xMan_OilON_Fdbk_H5 : Bool;   // Head#x manual oil feedback ON {x|x|x|x|O} / Head #5 manual oil feedback ON {x|x|x|x|O}
            xMan_FireON_Fdbk_H6 : Bool;   // Head#x manual fire ON Feeback {x|x|x|x|O} / Head #6 manual fire ON Feeback {x|x|x|x|O}
            xMan_FireOFF_Fdbk_H6 : Bool;   // Head#x manual fire OFF Feedback {x|x|x|x|O} / Head #6 manual fire OFF Feedback {x|x|x|x|O}
            xMan_OilON_Fdbk_H6 : Bool;   // Head#x manual oil feedback ON {x|x|x|x|O} / Head #6 manual oil feedback ON {x|x|x|x|O}
            xMan_FireON_Fdbk_H7 : Bool;   // Head#x manual fire ON Feeback {x|x|x|x|O} / Head #7 manual fire ON Feeback {x|x|x|x|O}
            xMan_FireOFF_Fdbk_H7 : Bool;   // Head#x manual fire OFF Feedback {x|x|x|x|O} / Head #7 manual fire OFF Feedback {x|x|x|x|O}
            xMan_OilON_Fdbk_H7 : Bool;   // Head#x manual oil feedback ON {x|x|x|x|O} / Head #7 manual oil feedback ON {x|x|x|x|O}
            xMan_FireON_Fdbk_H8 : Bool;   // Head#x manual fire ON Feeback {x|x|x|x|O} / Head #8 manual fire ON Feeback {x|x|x|x|O}
            xMan_FireOFF_Fdbk_H8 : Bool;   // Head#x manual fire OFF Feedback {x|x|x|x|O} / Head #8 manual fire OFF Feedback {x|x|x|x|O}
            xMan_OilON_Fdbk_H8 : Bool;   // Head#x manual oil feedback ON {x|x|x|x|O} / Head #8 manual oil feedback ON {x|x|x|x|O}
            xSpare24 : Bool;
            xSpare25 : Bool;
            xSpare26 : Bool;
            xSpare27 : Bool;
            xSpare28 : Bool;
            xSpare29 : Bool;
            xSpare30 : Bool;
            xSpare31 : Bool;
         END_STRUCT;
      END_STRUCT;
      tHMW : Struct   // HMI Write
         xResetUsageCounter_H1 : Bool;   // Head#x reset head usage counter {x|x|x|x|O} / Head #1 reset head usage counter {x|x|x|x|O}
         xResetUsageCounter_H2 : Bool := FALSE;   // Automatic mode request {x|x|x|x|O} / Head #2 reset head usage counter {x|x|x|x|O}
         xResetUsageCounter_H3 : Bool := FALSE;   // Manual mode request {x|x|x|x|O} / Head #3 reset head usage counter {x|x|x|x|O}
         xResetUsageCounter_H4 : Bool := FALSE;   // Bridge out of production request {x|x|x|x|O} / Head #4 reset head usage counter {x|x|x|x|O}
         xResetUsageCounter_H5 : Bool := FALSE;   // Bridge in production request {x|x|x|x|O} / Head #5 reset head usage counter {x|x|x|x|O}
         xResetUsageCounter_H6 : Bool := FALSE;   // Cut during glass break {x|x|x|x|O} / Head #6 reset head usage counter {x|x|x|x|O}
         xResetUsageCounter_H7 : Bool := FALSE;   // Motors and cards initialize {x|x|x|x|M} / Head #7 reset head usage counter {x|x|x|x|O}
         xResetUsageCounter_H8 : Bool := FALSE;   // Force the homing of the heads {x|x|x|x|M} / Head #8 reset head usage counter {x|x|x|x|O}
         xSpare8 : Bool := FALSE;   // Bridge offset calibration request {x|x|x|x|M}
         xSpare9 : Bool;
         xSpare10 : Bool;
         xSpare11 : Bool;
         xSpare12 : Bool;
         xSpare13 : Bool;
         xSpare14 : Bool := FALSE;
         xSpare15 : Bool := FALSE;
         xSpare16 : Bool := TRUE;
         xSpare17 : Bool := TRUE;
         xSpare18 : Bool := TRUE;
         xSpare19 : Bool := TRUE;
         xSpare20 : Bool := TRUE;
         xSpare21 : Bool := TRUE;
         xSpare22 : Bool := TRUE;
         xSpare23 : Bool := TRUE;
         xSpare24 : Bool;
         xSpare25 : Bool;
         xSpare26 : Bool;
         xSpare27 : Bool;
         xSpare28 : Bool;
         xSpare29 : Bool;
         xSpare30 : Bool;
         xSpare31 : Bool;
         xSpare : Array[0..15] of Bool;
         iSpare0 : Int;
         iSpare1 : Int;
         iSpare2 : Int;
         iSpare3 : Int;
         iSpare4 : Int;
         iSpare5 : Int;
         iSpare6 : Int;
         iSpare7 : Int;
         iSpare8 : Int;
         iSpare9 : Int;
         iSpare10 : Int;
         iSpare11 : Int;
         iSpare12 : Int;
         iSpare13 : Int;
         iSpare14 : Int;
         iSpare15 : Int;
         iSpare16 : Int := 0;
         dHeadFireONReaction_ms_H1 : DInt;   // Head#x fire ON reaction time [ms] {ms|s|0|1|M} / Head #1 fire ON reaction time [ms] {ms|s|0|1|M}
         dHeadFireOFFReaction_ms_H1 : DInt;   // Head#x fire OFF reaction time [ms] {ms|s|0|1|M} / Head #1 fire OFF reaction time [ms] {ms|s|0|1|M}
         dHeadOilONDelay_ms_H1 : DInt;   // Head#x Oil ON delay [ms]{ms|s|-2|2|O} / Head #1 Oil ON delay [ms]{ms|s|-2|2|O}
         dHeadOilOFFDelay_ms_H1 : DInt;   // Head#x Oil OFF delay [ms]{ms|s|-2|2|O} / Head #1 Oil OFF delay [ms]{ms|s|-2|2|O}
         dHeadFireONDelay_cmm_H1 : DInt;   // Head#x fire ON delay [mm/100] {mm/100|mm|-50|50|O} / Head #1 fire ON delay [mm/100] {mm/100|mm|-50|50|O}
         dHeadFireOFFDelay_cmm_H1 : DInt;   // Head#x fire OFF delay [mm/100] {mm/100|mm|-50|50|O} / Head #1 fire OFF delay [mm/100] {mm/100|mm|-50|50|O}
         dHeadPressure_mN_H1 : DInt;   // Head#x pressure value [N/1000] {N/1000|N|16|180|O} / Head #1 pressure value [N/1000] {N/1000|N|16|180|O}
         dHeadFireONReaction_ms_H2 : DInt;   // Head#x fire ON reaction time [ms] {ms|s|0|1|M} / Head #2 fire ON reaction time [ms] {ms|s|0|1|M}
         dHeadFireOFFReaction_ms_H2 : DInt;   // Head#x fire OFF reaction time [ms] {ms|s|0|1|M} / Head #2 fire OFF reaction time [ms] {ms|s|0|1|M}
         dHeadOilONDelay_ms_H2 : DInt;   // Head#x Oil ON delay [ms]{ms|s|-2|2|O} / Head #2 Oil ON delay [ms]{ms|s|-2|2|O}
         dHeadOilOFFDelay_ms_H2 : DInt;   // Head#x Oil OFF delay [ms]{ms|s|-2|2|O} / Head #2 Oil OFF delay [ms]{ms|s|-2|2|O}
         dHeadFireONDelay_cmm_H2 : DInt;   // Head#x fire ON delay [mm/100] {mm/100|mm|-50|50|O} / Head #2 fire ON delay [mm/100] {mm/100|mm|-50|50|O}
         dHeadFireOFFDelay_cmm_H2 : DInt;   // Head#x fire OFF delay [mm/100] {mm/100|mm|-50|50|O} / Head #2 fire OFF delay [mm/100] {mm/100|mm|-50|50|O}
         dHeadPressure_mN_H2 : DInt;   // Head#x pressure value [N/1000] {N/1000|N|16|180|O} / Head #2 pressure value [N/1000] {N/1000|N|16|180|O}
         dHeadFireONReaction_ms_H3 : DInt;   // Head#x fire ON reaction time [ms] {ms|s|0|1|M} / Head #3 fire ON reaction time [ms] {ms|s|0|1|M}
         dHeadFireOFFReaction_ms_H3 : DInt;   // Head#x fire OFF reaction time [ms] {ms|s|0|1|M} / Head #3 fire OFF reaction time [ms] {ms|s|0|1|M}
         dHeadOilONDelay_ms_H3 : DInt;   // Head#x Oil ON delay [ms]{ms|s|-2|2|O} / Head #3 Oil ON delay [ms]{ms|s|-2|2|O}
         dHeadOilOFFDelay_ms_H3 : DInt;   // Head#x Oil OFF delay [ms]{ms|s|-2|2|O} / Head #3 Oil OFF delay [ms]{ms|s|-2|2|O}
         dHeadFireONDelay_cmm_H3 : DInt;   // Head#x fire ON delay [mm/100] {mm/100|mm|-50|50|O} / Head #3 fire ON delay [mm/100] {mm/100|mm|-50|50|O}
         dHeadFireOFFDelay_cmm_H3 : DInt;   // Head#x fire OFF delay [mm/100] {mm/100|mm|-50|50|O} / Head #3 fire OFF delay [mm/100] {mm/100|mm|-50|50|O}
         dHeadPressure_mN_H3 : DInt;   // Head#x pressure value [N/1000] {N/1000|N|16|180|O} / Head #3 pressure value [N/1000] {N/1000|N|16|180|O}
         dHeadFireONReaction_ms_H4 : DInt;   // Head#x fire ON reaction time [ms] {ms|s|0|1|M} / Head #4 fire ON reaction time [ms] {ms|s|0|1|M}
         dHeadFireOFFReaction_ms_H4 : DInt;   // Head#x fire OFF reaction time [ms] {ms|s|0|1|M} / Head #4 fire OFF reaction time [ms] {ms|s|0|1|M}
         dHeadOilONDelay_ms_H4 : DInt;   // Head#x Oil ON delay [ms]{ms|s|-2|2|O} / Head #4 Oil ON delay [ms]{ms|s|-2|2|O}
         dHeadOilOFFDelay_ms_H4 : DInt;   // Head#x Oil OFF delay [ms]{ms|s|-2|2|O} / Head #4 Oil OFF delay [ms]{ms|s|-2|2|O}
         dHeadFireONDelay_cmm_H4 : DInt;   // Head#x fire ON delay [mm/100] {mm/100|mm|-50|50|O} / Head #4 fire ON delay [mm/100] {mm/100|mm|-50|50|O}
         dHeadFireOFFDelay_cmm_H4 : DInt;   // Head#x fire OFF delay [mm/100] {mm/100|mm|-50|50|O} / Head #4 fire OFF delay [mm/100] {mm/100|mm|-50|50|O}
         dHeadPressure_mN_H4 : DInt;   // Head#x pressure value [N/1000] {N/1000|N|16|180|O} / Head #4 pressure value [N/1000] {N/1000|N|16|180|O}
         dHeadFireONReaction_ms_H5 : DInt;   // Head#x fire ON reaction time [ms] {ms|s|0|1|M} / Head #5 fire ON reaction time [ms] {ms|s|0|1|M}
         dHeadFireOFFReaction_ms_H5 : DInt;   // Head#x fire OFF reaction time [ms] {ms|s|0|1|M} / Head #5 fire OFF reaction time [ms] {ms|s|0|1|M}
         dHeadOilONDelay_ms_H5 : DInt;   // Head#x Oil ON delay [ms]{ms|s|-2|2|O} / Head #5 Oil ON delay [ms]{ms|s|-2|2|O}
         dHeadOilOFFDelay_ms_H5 : DInt;   // Head#x Oil OFF delay [ms]{ms|s|-2|2|O} / Head #5 Oil OFF delay [ms]{ms|s|-2|2|O}
         dHeadFireONDelay_cmm_H5 : DInt;   // Head#x fire ON delay [mm/100] {mm/100|mm|-50|50|O} / Head #5 fire ON delay [mm/100] {mm/100|mm|-50|50|O}
         dHeadFireOFFDelay_cmm_H5 : DInt;   // Head#x fire OFF delay [mm/100] {mm/100|mm|-50|50|O} / Head #5 fire OFF delay [mm/100] {mm/100|mm|-50|50|O}
         dHeadPressure_mN_H5 : DInt;   // Head#x pressure value [N/1000] {N/1000|N|16|180|O} / Head #5 pressure value [N/1000] {N/1000|N|16|180|O}
         dHeadFireONReaction_ms_H6 : DInt;   // Head#x fire ON reaction time [ms] {ms|s|0|1|M} / Head #6 fire ON reaction time [ms] {ms|s|0|1|M}
         dHeadFireOFFReaction_ms_H6 : DInt;   // Head#x fire OFF reaction time [ms] {ms|s|0|1|M} / Head #6 fire OFF reaction time [ms] {ms|s|0|1|M}
         dHeadOilONDelay_ms_H6 : DInt;   // Head#x Oil ON delay [ms]{ms|s|-2|2|O} / Head #6 Oil ON delay [ms]{ms|s|-2|2|O}
         dHeadOilOFFDelay_ms_H6 : DInt;   // Head#x Oil OFF delay [ms]{ms|s|-2|2|O} / Head #6 Oil OFF delay [ms]{ms|s|-2|2|O}
         dHeadFireONDelay_cmm_H6 : DInt;   // Head#x fire ON delay [mm/100] {mm/100|mm|-50|50|O} / Head #6 fire ON delay [mm/100] {mm/100|mm|-50|50|O}
         dHeadFireOFFDelay_cmm_H6 : DInt;   // Head#x fire OFF delay [mm/100] {mm/100|mm|-50|50|O} / Head #6 fire OFF delay [mm/100] {mm/100|mm|-50|50|O}
         dHeadPressure_mN_H6 : DInt;   // Head#x pressure value [N/1000] {N/1000|N|16|180|O} / Head #6 pressure value [N/1000] {N/1000|N|16|180|O}
         dHeadFireONReaction_ms_H7 : DInt;   // Head#x fire ON reaction time [ms] {ms|s|0|1|M} / Head #7 fire ON reaction time [ms] {ms|s|0|1|M}
         dHeadFireOFFReaction_ms_H7 : DInt;   // Head#x fire OFF reaction time [ms] {ms|s|0|1|M} / Head #7 fire OFF reaction time [ms] {ms|s|0|1|M}
         dHeadOilONDelay_ms_H7 : DInt;   // Head#x Oil ON delay [ms]{ms|s|-2|2|O} / Head #7 Oil ON delay [ms]{ms|s|-2|2|O}
         dHeadOilOFFDelay_ms_H7 : DInt;   // Head#x Oil OFF delay [ms]{ms|s|-2|2|O} / Head #7 Oil OFF delay [ms]{ms|s|-2|2|O}